            xSpare13 : Bool;
            xSpare14 : Bool;
            xSpare15 : Bool;
            xSpare16 : Bool;
            xSpare17 : Bool;
            xSpare18 : Bool;
            xSpare19 : Bool;
            xSpare20 : Bool;
            xSpare21 : Bool;
            xSpare22 : Bool;
            xSpare23 : Bool;
            xSpare24 : Bool;
            xSpare25 : Bool;
            xSpare26 : Bool;
            xSpare27 : Bool;
            xSpare28 : Bool;
            xSpare29 : Bool;
            xSpare30 : Bool;
            xSpare31 : Bool;
         END_STRUCT;
      END_STRUCT;
   END_VAR
BEGIN
END_DATA_BLOCK

DATA_BLOCK "DB_Digitizer_2_HMI"   // DB2562
{ S7_Optimized_Access := 'FALSE' }
VERSION : 0.1
   VAR
      tALM : Struct   // HMI Alarms
         tE : Struct   // Emergency alarms
            xSpare_0 : Bool;
            xSpare_1 : Bool;
            xSpare_2 : Bool;
            xSpare_3 : Bool;
            xSpare_4 : Bool;
            xSpare_5 : Bool;
            xSpare_6 : Bool;
            xSpare_7 : Bool;
            xSpare_8 : Bool;
            xSpare_9 : Bool;
            xSpare_10 : Bool;
            xSpare_11 : Bool;
            xSpare_12 : Bool;
            xSpare_13 : Bool;
            xSpare_14 : Bool;
            xSpare_15 : Bool;
            xSpare_16 : Bool;
            xSpare_17 : Bool;
            xSpare_18 : Bool;
            xSpare_19 : Bool;
            xSpare_20 : Bool;
            xSpare_21 : Bool;
            xSpare_22 : Bool;
            xSpare_23 : Bool;
            xSpare_24 : Bool;
            xSpare_25 : Bool;
            xSpare_26 : Bool;
            xSpare_27 : Bool;
            xSpare_28 : Bool;
            xSpare_29 : Bool;
            xSpare_30 : Bool;
            xSpare_31 : Bool;
         END_STRUCT;
         tS : Struct   // Stopping faults
            xNoEncPulses : Bool;   // BQ.No encoder pulses
            xSpeedOutLimits : Bool;   // BQ.Speed outside min max limits
            xSpare_2 : Bool;
            xSpare_3 : Bool;
            xSpare_4 : Bool;
            xSpare_5 : Bool;
            xSpare_6 : Bool;
            xSpare_7 : Bool;
            xSpare_8 : Bool;
            xSpare_9 : Bool;
            xSpare_10 : Bool;
            xSpare_11 : Bool;
            xSpare_12 : Bool;
            xSpare_13 : Bool;
            xSpare_14 : Bool;
            xSpare_15 : Bool;
            xSpare_16 : Bool;
            xSpare_17 : Bool;
            xSpare_18 : Bool;
            xSpare_19 : Bool;
            xSpare_20 : Bool;
            xSpare_21 : Bool;
            xSpare_22 : Bool;
            xSpare_23 : Bool;
            xSpare_24 : Bool;
            xSpare_25 : Bool;
            xSpare_26 : Bool;
            xSpare_27 : Bool;
            xSpare_28 : Bool;
            xSpare_29 : Bool;
            xSpare_30 : Bool;
            xSpare_31 : Bool;
         END_STRUCT;
         tF : Struct   // Faults
            xMissingEncPulses : Bool;   // Missing encoder pulses
            xFm152SendError : Bool;   // FM152. Sending data error
            xFm152SendTimeout : Bool;   // FM152. Sending data timeout
            xFm152RecvTimeout : Bool;   // FM152.Receiving data timeout
            xSpare_4 : Bool;
            xSpare_5 : Bool;
            xSpare_6 : Bool;
            xSpare_7 : Bool;
            xSpare_8 : Bool;
            xSpare_9 : Bool;
            xSpare_10 : Bool;
            xSpare_11 : Bool;
            xSpare_12 : Bool;
            xSpare_13 : Bool;
            xSpare_14 : Bool;
            xSpare_15 : Bool;
            xSpare_16 : Bool;
            xSpare_17 : Bool;
            xSpare_18 : Bool;
            xSpare_19 : Bool;
            xSpare_20 : Bool;
            xSpare_21 : Bool;
            xSpare_22 : Bool;
            xSpare_23 : Bool;
            xSpare_24 : Bool;
            xSpare_25 : Bool;
            xSpare_26 : Bool;
            xSpare_27 : Bool;
            xSpare_28 : Bool;
            xSpare_29 : Bool;
            xSpare_30 : Bool;
            xSpare_31 : Bool;
         END_STRUCT;
         tW : Struct   // Warnings
            xSpare_0 : Bool;
            xSpare_1 : Bool;
            xSpare_2 : Bool;
            xSpare_3 : Bool;
            xSpare_4 : Bool;
            xSpare_5 : Bool;
            xSpare_6 : Bool;
            xSpare_7 : Bool;
            xSpare_8 : Bool;
            xSpare_9 : Bool;
            xSpare_10 : Bool;
            xSpare_11 : Bool;
            xSpare_12 : Bool;
            xSpare_13 : Bool;
            xSpare_14 : Bool;
            xSpare_15 : Bool;
            xSpare_16 : Bool;
            xSpare_17 : Bool;
            xSpare_18 : Bool;
            xSpare_19 : Bool;
            xSpare_20 : Bool;
            xSpare_21 : Bool;
            xSpare_22 : Bool;
            xSpare_23 : Bool;
            xSpare_24 : Bool;
            xSpare_25 : Bool;
            xSpare_26 : Bool;
            xSpare_27 : Bool;
            xSpare_28 : Bool;
            xSpare_29 : Bool;
            xSpare_30 : Bool;
            xSpare_31 : Bool;
         END_STRUCT;
      END_STRUCT;
      tHMR : Struct   // HMI Read
         xSpare0 : Bool;
         xSpare1 : Bool;
         xSpare2 : Bool;
         xSpare3 : Bool;
         xSpare4 : Bool;
         xSpare5 : Bool;
         xSpare6 : Bool;
         xSpare7 : Bool;
         xSpare8 : Bool;
         xSpare9 : Bool;
         xSpare10 : Bool;
         xSpare11 : Bool;
         xSpare12 : Bool;
         xSpare13 : Bool;
         xManualCommandEnabled : Bool;   // Manual Command enabled {x|x|x|x|O}
         xSpare15 : Bool;
         xSpare16 : Bool;
         xSpare17 : Bool;
         xSpare18 : Bool;
         xSpare19 : Bool;
         xSpare20 : Bool;
         xSpare21 : Bool;
         xSpare22 : Bool;
         xSpare23 : Bool;
         xSpare24 : Bool;
         xSpare25 : Bool;
         xSpare26 : Bool;
         xSpare27 : Bool;
         xSpare28 : Bool;
         xSpare29 : Bool;
         xSpare30 : Bool;
         xSpare31 : Bool;
         xSpare : Array[0..15] of Bool;
         iSpare0 : Int;
         iSpare1 : Int;
         iSpare2 : Int;
         iSpare3 : Int;
         iSpare4 : Int;
         iSpare5 : Int;
         iSpare6 : Int;
         iSpare7 : Int;
         iSpare8 : Int;
         iSpare9 : Int;
         iSpare10 : Int;
         iSpare11 : Int;
         iSpare12 : Int;
         iSpare13 : Int;
         iSpare14 : Int;
         iSpare15 : Int;
         iSpare16 : Int;
         dSpare0 : DInt;
         dEncoderStatus : DInt;   // Encoder status (1=Stop 3=Running 7=Anomaly)
         dFm152Status : DInt;   // Status of the Fm152 card
         dActualEncoderSpeed_mm_min : DInt;   // Actual encoder speed [mm/min]
         dCalibrationF1Unit_unit : DInt;   // Calibration actual F1 [unit]
         dCalibrationF2Unit_unit : DInt;   // Calibration actual F2 [unit]
         dCalibrationCardF1Unit_unit : DInt;   // Calibration actual F1 read from FM [unit]
         dCalibrationCardF2Unit_unit : DInt;   // Calibration actual F2 read from FM [unit]
         dSpare8 : DInt;
         dSpare9 : DInt;
         dSpare10 : DInt;
         dSpare11 : DInt;
         dSpare12 : DInt;
         dSpare13 : DInt;
         dSpare14 : DInt;
         dSpare15 : DInt;
         rSpare0 : Real;
         rSpare1 : Real;
         rSpare2 : Real;
         rSpare3 : Real;
         rSpare4 : Real;
         rSpare5 : Real;
         rSpare6 : Real;
         rSpare7 : Real;
         rSpare8 : Real;
         tManCmd : Struct
            xMan_DescEncFdbk : Bool;   // Manual mode. Feedback descent encoder
            xSpare1 : Bool;
            xSpare2 : Bool;
            xSpare3 : Bool;
            xSpare4 : Bool;
            xSpare5 : Bool;
            xSpare6 : Bool;
            xSpare7 : Bool;
            xSpare8 : Bool;
            xSpare9 : Bool;
            xSpare10 : Bool;
            xSpare11 : Bool;
            xSpare12 : Bool;
            xSpare13 : Bool;
            xSpare14 : Bool;
            xSpare15 : Bool;
            xSpare : Array[0..15] of Bool;
         END_STRUCT;
      END_STRUCT;
      tHMW : Struct   // HMI Write
         xCalibRequest : Bool;   // Calibration length request
         xCalibUpdateF1 : Bool;   // Calibration update F1 value
         xCalibUpdateF2 : Bool;   // Calibration update F2 value
         xGlassSensorEnabled : Bool;   // Glass presence sensor are enabled
         xSpare4 : Bool;
         xSpare5 : Bool;
         xSpare6 : Bool;
         xSpare7 : Bool;
         xSpare8 : Bool;
         xSpare9 : Bool;
         xSpare10 : Bool;
         xSpare11 : Bool;
         xSpare12 : Bool;
         xSpare13 : Bool;
         xEnableManualCommand : Bool;   // Enable Disable Manual command {x|x|x|x|O}
         xSpare15 : Bool;
         xSpare16 : Bool;
         xSpare17 : Bool;
         xSpare18 : Bool;
         xSpare19 : Bool;
         xSpare20 : Bool;
         xSpare21 : Bool;
         xSpare22 : Bool;
         xSpare23 : Bool;
         xSpare24 : Bool;
         xSpare25 : Bool;
         xSpare26 : Bool;
         xSpare27 : Bool;
         xSpare28 : Bool;
         xSpare29 : Bool;
         xSpare30 : Bool;
         xSpare31 : Bool;
         xSpare : Array[0..15] of Bool;
         iSpare0 : Int;
         iSpare1 : Int;
         iSpare2 : Int;
         iSpare3 : Int;
         iSpare4 : Int;
         iSpare5 : Int;
         iSpare6 : Int;
         iSpare7 : Int;
         iSpare8 : Int;
         iSpare9 : Int;
         iSpare10 : Int;
         iSpare11 : Int;
         iSpare12 : Int;
         iSpare13 : Int;
         iSpare14 : Int;
         iSpare15 : Int;
         iSpare16 : Int;
         dCalibTheoLength_cmm : DInt;   // Calibration theorical length [mm/100]
         dCalibWriteF2_unit : DInt;   // Calibration write F2 [unit]
         dCalibWriteF1_unit : DInt;   // Calibration write F1 [unit]
         dCalibRealLength_cmm : DInt;   // Calibration real length [mm/100]
         dRequestJogSpeed_mm_min : DInt;   // Jog speed requested [mm/min]
         dSpare5 : DInt;
         dSpare6 : DInt;
         dSpare7 : DInt;
         dSpare8 : DInt;
         dSpare9 : DInt;
         dSpare10 : DInt;
         dSpare11 : DInt;
         dSpare12 : DInt;
         dSpare13 : DInt;
         dSpare14 : DInt;
         dSpare15 : DInt;
         dSpare16 : DInt;
         rSpare0 : Real;
         rSpare1 : Real;
         rSpare2 : Real;
         rSpare3 : Real;
         rSpare4 : Real;
         rSpare5 : Real;
         rSpare6 : Real;
         rSpare7 : Real;
         rSpare8 : Real;
         tManCmd : Struct
            xMan_DescentEnc : Bool;   // Manual encoder descent
            xSpare1 : Bool;
            xSpare2 : Bool;
            xSpare3 : Bool;
            xSpare4 : Bool;
            xSpare5 : Bool;
            xSpare6 : Bool;
            xSpare7 : Bool;
            xSpare8 : Bool;
            xSpare9 : Bool;
            xSpare10 : Bool;
            xSpare11 : Bool;
            xSpare12 : Bool;
            xSpare13 : Bool;
            xSpare14 : Bool;
            xSpare15 : Bool;
            xSpare16 : Bool;
            xSpare17 : Bool;
            xSpare18 : Bool;
            xSpare19 : Bool;
            xSpare20 : Bool;
            xSpare21 : Bool;
            xSpare22 : Bool;
            xSpare23 : Bool;
            xSpare24 : Bool;
            xSpare25 : Bool;
            xSpare26 : Bool;
            xSpare27 : Bool;
            xSpare28 : Bool;
            xSpare29 : Bool;
            xSpare30 : Bool;
            xSpare31 : Bool;
         END_STRUCT;
      END_STRUCT;
   END_VAR
BEGIN
END_DATA_BLOCK

// folder: TaskErrors

DATA_BLOCK "RALRM_AUX_DB"   // DB59
{ S7_Optimized_Access := 'TRUE' }
VERSION : 0.1
   VAR RETAIN
      tAlm : Struct   // HMI Alarms
         tS : Struct   // Stopping faults
            xSpare_0 : Bool := FALSE;
            xSpare_1 : Bool := FALSE;
            xSpare_2 : Bool := FALSE;
            xSpare_3 : Bool := FALSE;
            xSpare_4 : Bool := FALSE;
            xSpare_5 : Bool := FALSE;
            xSpare_6 : Bool := FALSE;
            xSpare_7 : Bool := FALSE;
            xSpare_8 : Bool := FALSE;
            xSpare_9 : Bool := FALSE;
            xSpare_10 : Bool := FALSE;
            xSpare_11 : Bool := FALSE;
            xSpare_12 : Bool := FALSE;
            xSpare_13 : Bool := FALSE;
            xSpare_14 : Bool := FALSE;
            xSpare_15 : Bool := FALSE;
            xSpare_16 : Bool := FALSE;
            xSpare_17 : Bool := FALSE;
            xSpare_18 : Bool := FALSE;
            xSpare_19 : Bool := FALSE;
            xSpare_20 : Bool := FALSE;
            xSpare_21 : Bool := FALSE;
            xSpare_22 : Bool := FALSE;
            xSpare_23 : Bool := FALSE;
            xSpare_24 : Bool := FALSE;
            xSpare_25 : Bool := FALSE;
            xSpare_26 : Bool := FALSE;
            xSpare_27 : Bool := FALSE;
            xSpare_28 : Bool := FALSE;
            xSpare_29 : Bool := FALSE;
            xSpare_30 : Bool := FALSE;
            xSpare_31 : Bool := FALSE;
         END_STRUCT;
         tF : Struct   // Faults
            xDevice1 : Bool := FALSE;   // R13QF1.R13QF2.Power failure 230v auxiliary / Status device error.Device#1
            xDevice2 : Bool := FALSE;   // R18QF3.Power supply 24v logic / Status device error.Device#2
            xDevice3 : Bool := FALSE;   // R18QF4.Power supply 24v logic / Status device error.Device#3
            xDevice4 : Bool := FALSE;   // R18AP1.Redundancy 24v ok / Status device error.Device#4
            xDevice5 : Bool := FALSE;   // Status device error.Device#5
            xDevice6 : Bool := FALSE;   // Status device error.Device#6
            xDevice7 : Bool := FALSE;   // Status device error.Device#7
            xDevice8 : Bool := FALSE;   // Status device error.Device#8
            xDevice9 : Bool := FALSE;   // Status device error.Device#9
            xDevice10 : Bool := FALSE;   // Status device error.Device#10
            xSpare_10 : Bool := FALSE;
            xSpare_11 : Bool := FALSE;
            xSpare_12 : Bool;
            xSpare_13 : Bool;   // M250.R12KM1.Feedback rotation
            xSpare_14 : Bool;
            xSpare_15 : Bool;
            xSpare_16 : Bool;
            xSpare_17 : Bool;   // R204SP1.Compressed air presence cutting bridges
            xSpare_18 : Bool;
            xSpare_19 : Bool;
            xSpare_20 : Bool := FALSE;
            xSpare_21 : Bool := FALSE;
            xSpare_22 : Bool := FALSE;
            xSpare_23 : Bool := FALSE;
            xSpare_24 : Bool := FALSE;
            xSpare_25 : Bool := FALSE;
            xSpare_26 : Bool := FALSE;
            xSpare_27 : Bool := FALSE;
            xSpare_28 : Bool := FALSE;
            xSpare_29 : Bool := FALSE;
            xSpare_30 : Bool := FALSE;
            xSpare_31 : Bool := FALSE;
         END_STRUCT;
         tW : Struct   // Warnings
            xSpare_0 : Bool := FALSE;
            xSpare_1 : Bool := FALSE;
            xSpare_2 : Bool := FALSE;
            xSpare_3 : Bool := FALSE;
            xSpare_4 : Bool := FALSE;
            xSpare_5 : Bool := FALSE;
            xSpare_6 : Bool := FALSE;
            xSpare_7 : Bool := FALSE;
            xSpare_8 : Bool := FALSE;
            xSpare_9 : Bool := FALSE;
            xSpare_10 : Bool := FALSE;
            xSpare_11 : Bool := FALSE;
            xSpare_12 : Bool := FALSE;
            xSpare_13 : Bool := FALSE;
            xSpare_14 : Bool := FALSE;
            xSpare_15 : Bool := FALSE;
            xSpare_16 : Bool := FALSE;
            xSpare_17 : Bool := FALSE;
            xSpare_18 : Bool := FALSE;
            xSpare_19 : Bool := FALSE;
            xSpare_20 : Bool := FALSE;
            xSpare_21 : Bool := FALSE;
            xSpare_22 : Bool := FALSE;
            xSpare_23 : Bool := FALSE;
            xSpare_24 : Bool := FALSE;
            xSpare_25 : Bool := FALSE;
            xSpare_26 : Bool := FALSE;
            xSpare_27 : Bool := FALSE;
            xSpare_28 : Bool := FALSE;
            xSpare_29 : Bool := FALSE;
            xSpare_30 : Bool := FALSE;
            xSpare_31 : Bool := FALSE;
         END_STRUCT;
      END_STRUCT;
   END_VAR
BEGIN
END_DATA_BLOCK

// folder: TaskFast

DATA_BLOCK "FB_TrackDefects_V1_00_IDB"   // DB1
{ S7_Optimized_Access := 'TRUE' }
VERSION : 0.1
// stored: InstanceOfName FB_TrackDefects_V1.00
"FB_TrackDefects_V1.00"
BEGIN
END_DATA_BLOCK

DATA_BLOCK "DB_Defects"   // DB2
TITLE = Container of defect in extended mode
{ S7_Optimized_Access := 'TRUE' }
AUTHOR : A.Cigliutti
VERSION : 1.0
// Container of the defect in extended mode. These defect will be sent to optimizer and reporting system.
   VAR
      THIS : "UDT_DefectData_Tracking_Ext";
   END_VAR
BEGIN
END_DATA_BLOCK

DATA_BLOCK "FB_TrackCaps_V1_00_IDB"   // DB3
{ S7_Optimized_Access := 'TRUE' }
VERSION : 0.1
// stored: InstanceOfName FB_TrackCaps_V1.00
"FB_TrackCaps_V1.00"
BEGIN
END_DATA_BLOCK

DATA_BLOCK "FB_TrackEncoder_V1_00_IDB"   // DB4
{ S7_Optimized_Access := 'TRUE' }
VERSION : 0.1
// stored: InstanceOfName FB_TrackEncoder_V1.00
"FB_TrackEncoder_V1.00"
BEGIN
   IN_xSimulationActive := TRUE;
   IN_dSimulSpeed_mm_min := 10000;
   OUT_tHSCCount.loadValue0 := 16#0000_0000;
   OUT_tHSCCount.loadValue1 := 16#0000_0000;
   STC_AUX_tOutHSC.loadValue0 := 16#038D_6C80;
   STC_AUX_tOutHSC.loadValue1 := 16#0000_0000;
   STC_AUX_tOutHSC.swGate := TRUE;
   STC_AUX_tOutHSC.tmCtrlDQ0 := TRUE;
   STC_AUX_tOutHSC.tmCtrlDQ1 := TRUE;
   STC_ST_xCardInitialized := TRUE;
   STC_AUX_dNextMeterValue_cmm := 59600000;
   STC_AUX_dLastMeterValue_cmm := 59500000;
   STC_AUX_dMeterValueSent_cmm := 59600000;
   STC_AUX_lrTimingCounter_s := 4.59971222222222;
   STC_AUX_lrTimingCounterFast_s := 0.215018608888889;
   STC_AUX_lrElapsedTime_s := 0.00499898222222222;
   STC_AUX_lrRuntimeMemory_s := 16#0000_02A8_239A_5B38;
   STC_AUX_dLastCounterValue_cmm := 59518579;
   STC_AUX_dLastCounterValueFast_cmm := 59591502;
END_DATA_BLOCK

DATA_BLOCK "DB_Encoder"   // DB5
{ S7_Optimized_Access := 'TRUE' }
VERSION : 0.1
BEGIN
END_DATA_BLOCK

DATA_BLOCK "DB_Plates"   // DB6
{ S7_Optimized_Access := 'TRUE' }
VERSION : 0.1
BEGIN
END_DATA_BLOCK

DATA_BLOCK "GP_OB_Initialize_Fast_IDB"   // DB8
{ S7_Optimized_Access := 'TRUE' }
AUTHOR : Cigliutt
FAMILY : GP
VERSION : 1.1
// stored: InstanceOfName GP_OB_Initialize
"GP_OB_Initialize"
BEGIN
END_DATA_BLOCK

DATA_BLOCK "FB_Defects_Add_Fast_V1_00_IDB"   // DB14
{ S7_Optimized_Access := 'TRUE' }
VERSION : 0.1
// stored: InstanceOfName FB_Defects_Add_V1.00
"FB_Defects_Add_V1.00"
BEGIN
END_DATA_BLOCK

DATA_BLOCK "DB_RibbonData"   // DB40
{ S7_Optimized_Access := 'TRUE' }
VERSION : 0.1
BEGIN
END_DATA_BLOCK

DATA_BLOCK "FB_TrackRibbon_V1_00_IDB"   // DB41
{ S7_Optimized_Access := 'TRUE' }
VERSION : 0.1
// stored: InstanceOfName FB_TrackRibbon_V1.00
"FB_TrackRibbon_V1.00"
BEGIN
END_DATA_BLOCK

DATA_BLOCK "FB_CrossCutsModbusExchange_V1.00_DB"   // DB43
{ S7_Optimized_Access := 'TRUE' }
VERSION : 0.1
// stored: InstanceOfName FB_CrossCutsModbusExchange_V1.00
"FB_CrossCutsModbusExchange_V1.00"
BEGIN
END_DATA_BLOCK

DATA_BLOCK "FB_ISRASNAP_V1_00_IDB"   // DB53
{ S7_Optimized_Access := 'TRUE' }
VERSION : 0.1
// stored: InstanceOfName FB_ISRASNAP_V1.00
"FB_ISRASNAP_V1.00"
BEGIN
END_DATA_BLOCK

DATA_BLOCK "FB_CrossCut3ModbusExchange_V1.00_DB"   // DB64
{ S7_Optimized_Access := 'TRUE' }
VERSION : 0.1
// stored: InstanceOfName FB_CrossCutsModbusExchange_V1.00
"FB_CrossCutsModbusExchange_V1.00"
BEGIN
END_DATA_BLOCK

DATA_BLOCK "FB_CrossCut2ModbusExchange_V1.00_DB"   // DB65
{ S7_Optimized_Access := 'TRUE' }
VERSION : 0.1
// stored: InstanceOfName FB_CrossCutsModbusExchange_V1.00
"FB_CrossCutsModbusExchange_V1.00"
BEGIN
END_DATA_BLOCK

DATA_BLOCK "FB_CrossCut1ModbusExchange_V1.00_DB"   // DB66
{ S7_Optimized_Access := 'TRUE' }
VERSION : 0.1
// stored: InstanceOfName FB_CrossCutsModbusExchange_V1.00
"FB_CrossCutsModbusExchange_V1.00"
BEGIN
END_DATA_BLOCK

// folder: TaskMain

DATA_BLOCK "GP_OB_Initialize_Main_IDB"   // DB33
{ S7_Optimized_Access := 'TRUE' }
AUTHOR : Cigliutt
FAMILY : GP
VERSION : 1.1
// stored: InstanceOfName GP_OB_Initialize
"GP_OB_Initialize"
BEGIN
END_DATA_BLOCK

DATA_BLOCK "FB_BPSEthLink_ServerA_V1_00_IDB"   // DB34
{ S7_Optimized_Access := 'TRUE' }
VERSION : 0.1
// stored: InstanceOfName FB_BPSEthLink_V1.00
"FB_BPSEthLink_V1.00"
BEGIN
END_DATA_BLOCK

DATA_BLOCK "FB_Defects_Add_Main_V1_00_IDB"   // DB35
{ S7_Optimized_Access := 'TRUE' }
VERSION : 0.1
// stored: InstanceOfName FB_Defects_Add_V1.00
"FB_Defects_Add_V1.00"
BEGIN
END_DATA_BLOCK

DATA_BLOCK "FB_OptEthLink_V1_00_IDB"   // DB38
{ S7_Optimized_Access := 'TRUE' }
VERSION : 0.1
// stored: InstanceOfName FB_OptEthLink_V1.00
"FB_OptEthLink_V1.00"
BEGIN
END_DATA_BLOCK

DATA_BLOCK "FB_BPSEthLink_ServerB_V1_00_IDB"   // DB57
{ S7_Optimized_Access := 'TRUE' }
VERSION : 0.1
// stored: InstanceOfName FB_BPSEthLink_V1.00
"FB_BPSEthLink_V1.00"
BEGIN
END_DATA_BLOCK

DATA_BLOCK "DB_Z200_HMI"   // DB2011
{ S7_Optimized_Access := 'FALSE' }
VERSION : 0.1
   VAR
      tALM : Struct   // HMI Alarms
         tE : Struct   // Emergency alarms
            xSpare_0 : Bool := FALSE;
            xSpare_1 : Bool := FALSE;
            xSpare_2 : Bool := FALSE;
            xSpare_3 : Bool := FALSE;
            xSpare_4 : Bool := FALSE;
            xSpare_5 : Bool := FALSE;
            xSpare_6 : Bool := FALSE;
            xSpare_7 : Bool := FALSE;
            xSpare_8 : Bool := FALSE;
            xSpare_9 : Bool := FALSE;
            xSpare_10 : Bool := FALSE;
            xSpare_11 : Bool := FALSE;
            xSpare_12 : Bool := FALSE;
            xSpare_13 : Bool := FALSE;
            xSpare_14 : Bool := FALSE;
            xSpare_15 : Bool := FALSE;
            xSpare_16 : Bool := FALSE;
            xSpare_17 : Bool := FALSE;
            xSpare_18 : Bool := FALSE;
            xSpare_19 : Bool := FALSE;
            xSpare_20 : Bool := FALSE;
            xSpare_21 : Bool := FALSE;
            xSpare_22 : Bool := FALSE;
            xSpare_23 : Bool := FALSE;
            xSpare_24 : Bool := FALSE;
            xSpare_25 : Bool := FALSE;
            xSpare_26 : Bool := FALSE;
            xSpare_27 : Bool := FALSE;
            xSpare_28 : Bool := FALSE;
            xSpare_29 : Bool := FALSE;
            xSpare_30 : Bool := FALSE;
            xSpare_31 : Bool := FALSE;
         END_STRUCT;
         tS : Struct   // Stopping faults
            xSpare_0 : Bool := FALSE;
            xSpare_1 : Bool := FALSE;
            xSpare_2 : Bool := FALSE;
            xSpare_3 : Bool := FALSE;
            xSpare_4 : Bool := FALSE;
            xSpare_5 : Bool := FALSE;
            xSpare_6 : Bool := FALSE;
            xSpare_7 : Bool := FALSE;
            xSpare_8 : Bool := FALSE;
            xSpare_9 : Bool := FALSE;
            xSpare_10 : Bool := FALSE;
            xSpare_11 : Bool := FALSE;
            xSpare_12 : Bool := FALSE;
            xSpare_13 : Bool := FALSE;
            xSpare_14 : Bool := FALSE;
            xSpare_15 : Bool := FALSE;
            xSpare_16 : Bool := FALSE;
            xSpare_17 : Bool := FALSE;
            xSpare_18 : Bool := FALSE;
            xSpare_19 : Bool := FALSE;
            xSpare_20 : Bool := FALSE;
            xSpare_21 : Bool := FALSE;
            xSpare_22 : Bool := FALSE;
            xSpare_23 : Bool := FALSE;
            xSpare_24 : Bool := FALSE;
            xSpare_25 : Bool := FALSE;
            xSpare_26 : Bool := FALSE;
            xSpare_27 : Bool := FALSE;
            xSpare_28 : Bool := FALSE;
            xSpare_29 : Bool := FALSE;
            xSpare_30 : Bool := FALSE;
            xSpare_31 : Bool := FALSE;
         END_STRUCT;
         tF : Struct   // Faults
            xSpare_0 : Bool := TRUE;
            xProtectionCommandsAnomalies : Bool := FALSE;   // R18QF3.Power supply 24v logic
            xProtectionInternalInputAnomalies : Bool := FALSE;   // R18QF4.Power supply 24v logic
            xRedundancy24vOK1 : Bool := FALSE;   // R18AP1.Redundancy 24v ok
            xProtectionInternalOutputAnomalies : Bool := FALSE;   // R18QF7.Power supply 24v logic
            xProtectionExternalInputAnomalies : Bool := FALSE;   // R18QF8.Power supply 24v logic
            xSpare_6 : Bool := FALSE;
            xSpare_7 : Bool := FALSE;
            xSpare_8 : Bool := FALSE;
            xSpare_9 : Bool := FALSE;
            xSpare_10 : Bool := FALSE;
            xSpare_11 : Bool := FALSE;
            xSpare_12 : Bool;
            xSpare_13 : Bool;   // M250.R12KM1.Feedback rotation
            xSpare_14 : Bool;
            xSpare_15 : Bool;
            xSpare_16 : Bool;
            xCompressedAirCutting : Bool;   // R427SP1.Compressed air presence cutting bridges / R204SP1.Compressed air presence cutting bridges
            xPowerSupply24v_R18QF5_CPU_A : Bool;   // R18QF5.Power supply 24v CPU A
            xPowerSupply24v_R18QF6_CPU_B : Bool;   // R18QF6.Power supply 24v CPU B
            xPowerSupply24vProt1 : Bool := FALSE;
            xPowerSupply24vProt2 : Bool := FALSE;
            xMissingCPU_A_abilitation : Bool := FALSE;
            xMissingCPU_B_abilitation : Bool := FALSE;
            xSpare_24 : Bool := FALSE;
            xSpare_25 : Bool := FALSE;
            xSpare_26 : Bool := FALSE;
            xSpare_27 : Bool := FALSE;
            xSpare_28 : Bool := FALSE;
            xSpare_29 : Bool := FALSE;
            xSpare_30 : Bool := FALSE;
            xSpare_31 : Bool := FALSE;
         END_STRUCT;
         tW : Struct   // Warnings
            xPowerFailure230vAux : Bool := FALSE;   // R11QF2/3.Power failure 230v auxiliary
            xSpare_1 : Bool := FALSE;
            xSpare_2 : Bool := FALSE;
            xSpare_3 : Bool := FALSE;
            xSpare_4 : Bool := FALSE;
            xSpare_5 : Bool := FALSE;
            xSpare_6 : Bool := FALSE;
            xSpare_7 : Bool := FALSE;
            xSpare_8 : Bool := FALSE;
            xSpare_9 : Bool := FALSE;
            xSpare_10 : Bool := FALSE;
            xSpare_11 : Bool := FALSE;
            xSpare_12 : Bool := FALSE;
            xSpare_13 : Bool := FALSE;
            xSpare_14 : Bool := FALSE;
            xSpare_15 : Bool := FALSE;
            xSpare_16 : Bool := FALSE;
            xSpare_17 : Bool := FALSE;
            xSpare_18 : Bool := FALSE;
            xSpare_19 : Bool := FALSE;
            xSpare_20 : Bool := FALSE;
            xSpare_21 : Bool := FALSE;
            xSpare_22 : Bool := FALSE;
            xSpare_23 : Bool := FALSE;
            xSpare_24 : Bool := FALSE;
            xSpare_25 : Bool := FALSE;
            xSpare_26 : Bool := FALSE;
            xSpare_27 : Bool := FALSE;
            xSpare_28 : Bool := FALSE;
            xSpare_29 : Bool := FALSE;
            xSpare_30 : Bool := FALSE;
            xSpare_31 : Bool := FALSE;
         END_STRUCT;
      END_STRUCT;
      tHMR : Struct   // HMI Read
         xSpare0 : Bool;
         xSpare1 : Bool;
         xSpare2 : Bool;
         xSpare3 : Bool;
         xSpare4 : Bool;
         xSpare5 : Bool;
         xSpare6 : Bool;
         xSpare7 : Bool;
         xSpare8 : Bool;
         xSpare9 : Bool;
         xSpare10 : Bool;
         xSpare11 : Bool;
         xSpare12 : Bool;
         xSpare13 : Bool;
         xSpare14 : Bool;
         xZoneAlarm : Bool := FALSE;   // Zone alarm {X|X|X|X|O}
         xSpare16 : Bool;
         xSpare17 : Bool;
         xSpare18 : Bool;
         xSpare19 : Bool;
         xSpare20 : Bool;
         xSpare21 : Bool;
         xSpare22 : Bool;
         xSpare23 : Bool;
         xSpare24 : Bool;
         xSpare25 : Bool;
         xSpare26 : Bool;
         xSpare27 : Bool;
         xSpare28 : Bool;
         xSpare29 : Bool;
         xSpare30 : Bool;
         xSpare31 : Bool;
         xSpare : Array[0..15] of Bool;
         iSpare0 : Int;
         iSpare1 : Int;
         iSpare2 : Int;
         iSpare3 : Int;
         iSpare4 : Int;
         iSpare5 : Int;
         iSpare6 : Int;
         iSpare7 : Int;
         iSpare8 : Int;
         iSpare9 : Int;
         iSpare10 : Int;
         iSpare11 : Int;
         iSpare12 : Int;
         iSpare13 : Int;
         iSpare14 : Int;
         iSpare15 : Int;
         iSpare16 : Int;
         dSpare0 : DInt;
         dZoneState : DInt := 1024;   // Zone status (1=CycleON 2=StopCyc 4=CycleReq 8=StopReq 1024=E-Stop) {X|X|X|X|O}
         dCabinetStatusMCC1200 : DInt := 1;   // Cabinet status MCC1200 (0=OK;1=General power alarm;2=Local power alarm) {X|X|X|X|O}
         dSpare3 : DInt;
         dSpare4 : DInt;
         dSpare5 : DInt;
         dSpare6 : DInt;
         dSpare7 : DInt;
         dSpare8 : DInt;
         dSpare9 : DInt;
         dSpare10 : DInt;
         dSpare11 : DInt;
         dSpare12 : DInt;
         dSpare13 : DInt;
         dSpare14 : DInt;
         dSpare15 : DInt;
         rSpare0 : Real;
         rSpare1 : Real;
         rSpare2 : Real;
         rSpare3 : Real;
         rSpare4 : Real;
         rSpare5 : Real;
         rSpare6 : Real;
         rSpare7 : Real;
         rSpare8 : Real;
         tManCmd : Struct
            xSpare0 : Bool;
            xSpare1 : Bool;
            xSpare2 : Bool;
            xSpare3 : Bool;
            xSpare4 : Bool;
            xSpare5 : Bool;
            xSpare6 : Bool;
            xSpare7 : Bool;
            xSpare8 : Bool;
            xSpare9 : Bool;
            xSpare10 : Bool;
            xSpare11 : Bool;
            xSpare12 : Bool;
            xSpare13 : Bool;
            xSpare14 : Bool;
            xSpare15 : Bool;
            xSpare : Array[0..15] of Bool;
         END_STRUCT;
      END_STRUCT;
      tHMW : Struct   // HMI Write
         xSpare0 : Bool;
         xSpare1 : Bool;
         xSpare2 : Bool;
         xSpare3 : Bool;
         xSpare4 : Bool;
         xSpare5 : Bool := FALSE;
         xSpare6 : Bool := FALSE;
         xSpare7 : Bool := FALSE;
         xSpare8 : Bool;
         xSpare9 : Bool;
         xSpare10 : Bool;
         xSpare11 : Bool;
         xSpare12 : Bool;
         xSpare13 : Bool;
         xSpare14 : Bool;
         xSpare15 : Bool := FALSE;
         xSpare16 : Bool := FALSE;
         xSpare17 : Bool;
         xSpare18 : Bool;
         xSpare19 : Bool;
         xSpare20 : Bool;
         xSpare21 : Bool;
         xSpare22 : Bool;
         xSpare23 : Bool;
         xSpare24 : Bool;
         xSpare25 : Bool;
         xSpare26 : Bool;
         xSpare27 : Bool;
         xSpare28 : Bool;
         xSpare29 : Bool;
         xSpare30 : Bool;
         xSpare31 : Bool;
         xSpare : Array[0..15] of Bool;
         iSpare0 : Int;
         iSpare1 : Int;
         iSpare2 : Int;
         iSpare3 : Int;
         iSpare4 : Int;
         iSpare5 : Int;
         iSpare6 : Int;
         iSpare7 : Int;
         iSpare8 : Int;
         iSpare9 : Int;
         iSpare10 : Int;
         iSpare11 : Int;
         iSpare12 : Int;
         iSpare13 : Int;
         iSpare14 : Int;
         iSpare15 : Int;
         iSpare16 : Int;
         dSpare0 : DInt;
         dSpare1 : DInt;
         dSpare2 : DInt;
         dSpare3 : DInt;
         dSpare4 : DInt;
         dSpare5 : DInt;
         dSpare6 : DInt;
         dSpare7 : DInt;
         dSpare8 : DInt;
         dSpare9 : DInt;
         dSpare10 : DInt;
         dSpare11 : DInt;
         dSpare12 : DInt;
         dSpare13 : DInt;
         dSpare14 : DInt;
         dSpare15 : DInt;
         dSpare16 : DInt;
         rSpare0 : Real;
         rSpare1 : Real;
         rSpare2 : Real;
         rSpare3 : Real;
         rSpare4 : Real;
         rSpare5 : Real;
         rSpare6 : Real;
         rSpare7 : Real;
         rSpare8 : Real;
         tManCmd : Struct
            xSpare0 : Bool;
            xSpare1 : Bool;
            xSpare2 : Bool;
            xSpare3 : Bool;
            xSpare4 : Bool;
            xSpare5 : Bool;
            xSpare6 : Bool;
            xSpare7 : Bool;
            xSpare8 : Bool;
            xSpare9 : Bool;
            xSpare10 : Bool;
            xSpare11 : Bool;
            xSpare12 : Bool;
            xSpare13 : Bool;
            xSpare14 : Bool;
            xSpare15 : Bool;
            xSpare16 : Bool;
            xSpare17 : Bool;
            xSpare18 : Bool;
            xSpare19 : Bool;
            xSpare20 : Bool;
            xSpare21 : Bool;
            xSpare22 : Bool;
            xSpare23 : Bool;
            xSpare24 : Bool;
            xSpare25 : Bool;
            xSpare26 : Bool;
            xSpare27 : Bool;
            xSpare28 : Bool;
            xSpare29 : Bool;
            xSpare30 : Bool;
            xSpare31 : Bool;
         END_STRUCT;
      END_STRUCT;
   END_VAR
BEGIN
END_DATA_BLOCK

// folder: TaskMain/Z201

DATA_BLOCK "Z201"   // DB18
{ S7_Optimized_Access := 'TRUE' }
VERSION : 0.1
   VAR
      tmOFF_ResetAlarm : "UDT_IECTOFF_V1.00";   // Reset alarm / Reset alarm retentive timer
      tmON_24Vdc : "UDT_IECTON_V1.00";   // Presence 24Vdc timer / 24VDC ok delayed timer
      tmON_EmergencyOK : "UDT_IECTON_V1.00";   // Emergency OK timer / Emergency ok delayed timer
      tmON_CycleOnDelayed : "UDT_IECTON_V1.00";   // Cycle ON delayed
      tmON_CycleOn : "UDT_IECTON_V1.00";   // Cycle ON timer
      tmOFF_GeneralReset : "UDT_IECTOFF_V1.00";   // General reset retentive timer
      ST_xZoneError : Bool := FALSE;   // Zone error / Zone is in error
      ST_xFaultsEnabled : Bool := FALSE;   // Faults enabled
      ST_xZoneEmergency : Bool := FALSE;   // Cumulative of emergency faults active / Zone is in emergency
      ST_xZoneFaults : Bool := FALSE;   // Cumulative of zone faults / Zone is in faults
      ST_xZoneStoppingFaults : Bool := FALSE;   // Cumulative of zone stopping faults / Zone is in stopping faults
      ST_xOutputEnabledM216Fan : Bool;   // Output enable M216 fan / Output enable M250 fan
      ST_xOutputEnabledM209Chips : Bool;   // Output enable M209 chips blower / Output enable M272 chips blower
      ST_xZoneWarnings : Bool := FALSE;   // Cumulative of zone warning / Zone is in warning
      ST_xCycleON : Bool := FALSE;   // Zone in cycle ON / Cycle ON
      ST_xConditionOKStopCycle : Bool := FALSE;   // Condition ok to accept stop cycle
      ST_xCycleONDelayed : Bool := FALSE;   // Cycle ON delayed
      ST_xConditionOkPhaseAdvancement : Bool := FALSE;   // Condition ok for phase advancement
      ST_xConditionOkCycleON : Bool := FALSE;   // Condition ok for cycle ON
      ST_xMachineReset : Bool := FALSE;   // Machine reset request
      ST_xPLC1 : Bool := TRUE;   // This is PLC 1
      ST_xPLC2 : Bool := FALSE;   // This is PLC 2
      ST_xThisPlcActive : Bool := TRUE;   // This PLC is active
      ST_xStartCycleRequest : Bool := FALSE;   // Request start cycle
      ST_xStopCycleRequest : Bool := FALSE;   // Request stop cycle
      ST_xM209GlassBreak : Bool;   // M209 Chips blower glass break / M272 Chips blower glass break
      ST_xAllarmOFF : Bool;
      OSR_xStartCycle : Bool := FALSE;   // OSR start cycle
      OSR_xStopCycle : Bool := FALSE;   // OSR stop cycle
      OSR_xForceStopCycle : Bool := FALSE;   // OSR force stop cycle
      OSR_xChipsBlowerON : Bool;   // OSR chips blower on
      OSR_xSBResetAnomaly : Bool;   // OSR reset anomaly
      OS_xStartCycle : Bool := FALSE;   // OS start cycle
      OS_xStopCycle : Bool := FALSE;   // OS stop cycle
      OS_xForceStopCycle : Bool := FALSE;   // OS force stop cycle
      OS_xChipsBlowerON : Bool;   // OS chips blower on
      OS_xCpuActive : Bool;   // OS Cpu active
      OSR_xCpuActive : Bool;   // OSR Cpu active
      ST_xStopCycleAccepted : Bool := FALSE;   // Stop cycle accepted
      AUX_tmON_M216FanFeedback : "UDT_IECTON_V1.00";   // M216 Fan feedback anomaly / M250 Fan feedback anomaly
      AUX_tmON_M209ChipsFeedback : "UDT_IECTON_V1.00";   // M209 Chips blower feedback anomaly / M272 Chips blower feedback anomaly
      tOutputs : Struct
         xPLC1On : Bool;   // o.A406AP1.A255HL4.EnableCPUA
         xPLC2On : Bool;   // o.A406AP1.A255HL5.EnableCPUB
         xRunFanM216 : Bool;   // Run fan
         xRunFanM209 : Bool;   // Run fan
         xEmergencyON : Bool;   // o.A406AP1.A255HL1/1A.EmergencyON
         xSafetiesON : Bool;   // o.A406AP1.A255HL3.SafetiesON
         xHLResetAnomaly : Bool;   // o.A406AP1.A207SB1.HLResetAnomalyZ200
         xHAAlarm : Bool;   // o.A401AP1.A416HA1.Alarm
         xHLchipBlowerM209On : Bool;   // o.A406AP1.HL ChipBlowerM209On
      END_STRUCT;
      tInputs : Struct
         xPowerSupply230vAux : Bool := FALSE;   // i.A406AP1.A10QF1/2.PowerFailure230VAuxiliary / i.R195AP1.R13QF1/2.PowerFailure230VAuxiliary
         xPowerSuppluyOut24vUnderUpsEmOk : Bool;   // i.R195AP1.R18AP1.Redundacy24VOk / i.A406AP1.A108QF5.Out24vUnderUpsEmOk
         xPowerSupply24vLogic1 : Bool := FALSE;   // i.A406AP1.A18QF3.PowerSupply24VLogic / i.R195AP1.R18QF3.PowerSupply24VLogic
         xPowerSupply24vLogic2 : Bool := FALSE;   // i.A406AP1.A18QF4.PowerSupply24VLogic / i.R195AP1.R18QF4.PowerSupply24VLogic
         xPowerSupply24vLogic3 : Bool := FALSE;   // i.A406AP1.A19QF1.PowerSupply24VLogic / i.R195AP1.R18QF4.PowerSupply24VLogic
         xPowerSupply24vLogic4 : Bool := FALSE;   // i.A406AP1.A19QF2.PowerSupply24VLogic / i.R195AP1.R18QF4.PowerSupply24VLogic
         xPowerSuppluyOut24vUnderEmOk : Bool;   // i.A406AP1.A108QF6.Out24vUnderUpsEmOk
         xPowerSupply24vDrive2 : Bool;   // i.A406AP1.A20QF4.PowerSupply24VDrive
         xMainEmergencyON : Bool := FALSE;   // i.A406AP1.A45KE1.MainEmergencyON / i.R195AP1.R18QF4.PowerSupply24VLogic
         xEmergencyONArea201 : Bool;   // i.A406AP1.EmergencyArea201ON
         xEmergencyONArea301 : Bool;   // i.A406AP1.EmergencyArea301ON
         xEmergencyONArea302 : Bool;   // i.A406AP1.EmergencyArea302ON
         xEmergencyONArea303 : Bool;   // i.A406AP1.F38KE1.EmergencyArea303ON
         xEmergencyONArea601 : Bool;   // i.A406AP1.A38KE2.EmergencyArea601ON
         xEmergencyONArea701 : Bool;   // i.A406AP1.A39KE1.EmergencyArea701ON
         xDriveSupply2 : Bool;   // i.A406AP1.A52QM1.DriveSupply
         xCPUAEnabled : Bool := FALSE;   // i.A151AP1.Selection CPU A / i.R150AP1.CPU A Enabled
         xCPUBEnabled : Bool := TRUE;   // i.A151AP1.Selection CPU B / i.R150AP1.CPU B Enabled
         xCPUARecognition : Bool := FALSE;   // i.A151AP1.Recognition CPU A / i.R150AP1.Recognition CPU A
         xCPUBRecognition : Bool := FALSE;   // i.A151AP1.Recognition CPU B / i.R150AP1.Recognition CPU B
         xM216FanProtection : Bool;   // i.A406AP1.A141QM1.ProtectionRotationM216 / i.R195AP1.R12KM1.FeedbackRotationM250
         xM216FanFeedback : Bool;   // i.A406AP1.A141KM1.FeedbackRotationM216 / i.R195AP1.R12KM1.FeedbackRotationM250
         xM209FanFeedback : Bool;   // i.A406AP1.A178KM1.FeedbackRotationM209 / i.R195AP1.R12KM1.FeedbackRotationM250
         xM209FanProtection : Bool;   // i.A406AP1.FanProtectionOnM209 / i.R195AP1.R12KM1.FeedbackRotationM250
         xEmLocMCC1201 : Bool;   // i.A406AP1.A118SB1.EmergencyLocalization_MCC1201
         xEmLocCS4201 : Bool;   // i.A406AP1.A33SB2.EmergencyLocalization_CS4201
         xEmLocM203 : Bool;   // i.A406AP1.M203_SB3.EmergencyLocalization_M203
         xEmLocM204S_1 : Bool;   // i.A406AP1.M204S_SB3.EmergencyLocalization_M203S
         xEmLocM204S_2 : Bool;   // i.A406AP1.M204S_SB4.EmergencyLocalization_M203S
         xEmLocM211_1 : Bool;   // i.A406AP1.M211SB1.EmergencyLocalization_M211
         xEmLocM211_2 : Bool;   // i.A406AP1.M211SB2.EmergencyLocalization_M211
         xEmLocM214_1 : Bool;   // i.A406AP1.M214SB1.EmergencyLocalization_M214
         xEmLocM214_2 : Bool;   // i.A406AP1.M214SB2.EmergencyLocalization_M214
         xEmLocM218_1 : Bool;   // i.A406AP1.M218SB1.EmergencyLocalization_M218
         xEmLocM218_2 : Bool;   // i.A406AP1.M218SB2.EmergencyLocalization_M218
         xEmLocCS4202 : Bool;   // i.A406AP1.CS4201SB2.EmergencyLocalization_CS4201
         xSBResetAnomalyZ200 : Bool;   // i.A406AP1.A207SB1.ResetAnomalyZ200
         xSBglassReqToQLT : Bool;   // i.CS4202.E406AP1.E547SB5.GlassRequestToQLT
         xSBchipBlowerON_M209 : Bool;   // i.A406AP1.M209SB1 ChipsBlower ON
      END_STRUCT;
   END_VAR
BEGIN
END_DATA_BLOCK

DATA_BLOCK "ZUPS"   // DB29
{ S7_Optimized_Access := 'TRUE' }
VERSION : 0.1
   VAR
      tmON_EmergencyUPSOK : "UDT_IECTON_V1.00";   // Emergency UPS ok delayed timer
      tmON_CycleOnDelayed : "UDT_IECTON_V1.00";   // Cycle ON delayed
      tmON_CycleOn : "UDT_IECTON_V1.00";   // Cycle ON timer
      tmOFF_ResetAlarm : "UDT_IECTOFF_V1.00";   // Reset alarm / Reset alarm retentive timer
      ST_xZoneError : Bool := FALSE;   // Zone error / Zone is in error
      ST_xFaultsEnabled : Bool := TRUE;   // Faults enabled
      ST_xZoneEmergency : Bool := TRUE;   // Cumulative of emergency faults active / Zone is in emergency
      ST_xZoneFaults : Bool := TRUE;   // Cumulative of zone faults / Zone is in faults
      ST_xZoneStoppingFaults : Bool := FALSE;   // Cumulative of zone stopping faults / Zone is in stopping faults
      ST_xZoneWarnings : Bool := FALSE;   // Cumulative of zone warning / Zone is in warning
      ST_xCycleON : Bool := TRUE;   // Zone in cycle ON / Cycle ON
      ST_xConditionOKStopCycle : Bool := TRUE;   // Condition ok to accept stop cycle
      ST_xCycleONDelayed : Bool := TRUE;   // Cycle ON delayed
      ST_xConditionOkPhaseAdvancement : Bool := FALSE;   // Condition ok for phase advancement
      ST_xConditionOkCycleON : Bool := FALSE;   // Condition ok for cycle ON
      ST_xStartCycleRequest : Bool := FALSE;   // Request start cycle
      ST_xStopCycleRequest : Bool := FALSE;   // Request stop cycle
      OSR_xStartCycle : Bool := FALSE;   // OSR start cycle
      OSR_xStopCycle : Bool := FALSE;   // OSR stop cycle
      OSR_xForceStopCycle : Bool := FALSE;   // OSR force stop cycle
      OSR_xChipsBlowerON : Bool;   // OSR chips blower on
      OS_xStartCycle : Bool := FALSE;   // OS start cycle
      OS_xStopCycle : Bool := FALSE;   // OS stop cycle
      OS_xForceStopCycle : Bool := FALSE;   // OS force stop cycle
      OS_xChipsBlowerON : Bool;   // OS chips blower on
      OS_xCpuActive : Bool;   // OS Cpu active
      OSR_xCpuActive : Bool;   // OSR Cpu active
      OSR_xSBResetAnomaly : Bool;   // OSR reset anomaly
      ST_xStopCycleAccepted : Bool := FALSE;   // Stop cycle accepted
      tOutputs : Struct
         xUPSEmergencyON : Bool;   // o.A195AP1.A255HL2.UPSEmergencyON
         xHAAlarm : Bool;   // o.A401AP1.A416HA1.Alarm
      END_STRUCT;
      tInputs : Struct
         xPowerSupply24vDrive1 : Bool;   // i.A406AP1.A110QF2.PowerSupply24VDrive
         xEmergencyONAreaUPS : Bool := FALSE;   // i.A406AP1.A117KE1.EmergencyAreaUPSON / i.R195AP1.R18QF4.PowerSupply24VLogic
         xDriveSupply1 : Bool;   // i.A406AP1.A51QM1.DriveSupply
         xUPSEmLocMCC1201 : Bool;   // i.A406AP1.A117SB1.EmergencyLocalizationUPS_MCC1201
         xUPSEmLocM204S_1 : Bool;   // i.A406AP1.M204S_SB1.EmergencyLocalizationUPS_M204S
         xUPSEmLocM204S_2 : Bool;   // i.A406AP1.M204S_SB2.EmergencyLocalizationUPS_M204S
         xUPSEmLocCS4201 : Bool;   // i.A406AP1.M204S_SB2.EmergencyLocalizationUPS_M204S
      END_STRUCT;
   END_VAR
BEGIN
END_DATA_BLOCK

DATA_BLOCK "FB_Z200Conveyor_M201_IDB"   // DB101
{ S7_Optimized_Access := 'TRUE' }
VERSION : 0.1
// stored: InstanceOfName FB_Z200Conveyor_SinamicsMotor
"FB_Z200Conveyor_SinamicsMotor"
BEGIN
END_DATA_BLOCK

DATA_BLOCK "FB_Z200Conveyor_M204_IDB"   // DB102
{ S7_Optimized_Access := 'TRUE' }
VERSION : 0.1
// stored: InstanceOfName FB_Z200Conveyor_SinamicsMotor
"FB_Z200Conveyor_SinamicsMotor"
BEGIN
END_DATA_BLOCK

DATA_BLOCK "FB_Z200Conveyor_M205_IDB"   // DB103
{ S7_Optimized_Access := 'TRUE' }
VERSION : 0.1
// stored: InstanceOfName FB_Z200Conveyor_SinamicsMotor
"FB_Z200Conveyor_SinamicsMotor"
BEGIN
END_DATA_BLOCK

DATA_BLOCK "FB_Z200Conveyor_M208_IDB"   // DB104
{ S7_Optimized_Access := 'TRUE' }
VERSION : 0.1
// stored: InstanceOfName FB_Z200Conveyor_SinamicsMotor
"FB_Z200Conveyor_SinamicsMotor"
BEGIN
END_DATA_BLOCK

DATA_BLOCK "FB_Z200Conveyor_M211_iDB"   // DB105
{ S7_Optimized_Access := 'TRUE' }
VERSION : 0.1
// stored: InstanceOfName FB_Z200Conveyor_SinamicsMotor
"FB_Z200Conveyor_SinamicsMotor"
BEGIN
END_DATA_BLOCK

DATA_BLOCK "FB_Z200Conveyor_M214_iDB"   // DB106
{ S7_Optimized_Access := 'TRUE' }
VERSION : 0.1
// stored: InstanceOfName FB_Z200Conveyor_SinamicsMotor
"FB_Z200Conveyor_SinamicsMotor"
BEGIN
END_DATA_BLOCK

DATA_BLOCK "FB_Z200Conveyor_M218_IDB"   // DB107
{ S7_Optimized_Access := 'TRUE' }
VERSION : 0.1
// stored: InstanceOfName FB_Z200Conveyor_SinamicsMotor
"FB_Z200Conveyor_SinamicsMotor"
BEGIN
END_DATA_BLOCK

DATA_BLOCK "FB_BreakerM206_V1_00_IDB"   // DB109
{ S7_Optimized_Access := 'TRUE' }
VERSION : 0.1
// stored: InstanceOfName FB_BreakerM206_V1.00
"FB_BreakerM206_V1.00"
BEGIN
END_DATA_BLOCK

DATA_BLOCK "FB_DropConveyor_IDB"   // DB110
{ S7_Optimized_Access := 'TRUE' }
VERSION : 0.1
// stored: InstanceOfName FB_DropConveyor
"FB_DropConveyor"
BEGIN
END_DATA_BLOCK

DATA_BLOCK "FB_IO_EmergencyCuttingBridge_DB"   // DB111
{ S7_Optimized_Access := 'TRUE' }
VERSION : 0.1
// stored: InstanceOfName FB_IO_EmergencyCuttingBridge
"FB_IO_EmergencyCuttingBridge"
BEGIN
END_DATA_BLOCK

DATA_BLOCK "CU_A250AP1_IDB"   // DB218
{ S7_Optimized_Access := 'FALSE' }
AUTHOR : Armitano
VERSION : 1.7
// stored: InstanceOfName SINAMICS_ControlUnit
"SINAMICS_ControlUnit"
BEGIN
END_DATA_BLOCK

DATA_BLOCK "CU_A260AP1_IDB"   // DB219
{ S7_Optimized_Access := 'FALSE' }
AUTHOR : Armitano
VERSION : 1.7
// stored: InstanceOfName SINAMICS_ControlUnit
"SINAMICS_ControlUnit"
BEGIN
END_DATA_BLOCK

